(* Logix 5000 project; controller FV vendor 1 type 14 code 217 rev 31.11; software revision 31.00; part 26 of 63 *)
(* tags used below, declared in another part *)
   Alarm_Reset : BOOL;
   CheckTimeMask : INT;
   comms_to_mc_write_enabled : BOOL;
   comms_to_mv_route_write_enabled : BOOL;
   Default_Check_Time : DINT;
   Delphi_Does_Eng_Func : BOOL;
   FR_B3 : INT[255];   // BINARY
   fr_comms_from_mv_route : MESSAGE;
   fr_comms_from_mvfv_cip : MESSAGE;
   fr_comms_to_MC : MESSAGE;
   fr_comms_to_MC_timer : TIMER;
   fr_comms_to_mv_route : MESSAGE;
   fr_comms_to_mv_route_timer : TIMER;
   FR_FV27_AV08 : PlantItem;   // FV27_AV08
   FR_FV28_AV08 : PlantItem;   // FV28_AV08
   FR_FV29_AV08 : PlantItem;   // FV29_AV08
   FR_FV30_AV08 : PlantItem;   // FV30_AV08
   FR_FV31_AV08 : PlantItem;   // FV31_AV08
   FR_FVR1_P01 : PlantItem;   // FVR1_P01
   FR_FVR1_P01_ALARM : ALARM_DIGITAL;
   FR_FVR1_P01_D : ALIAS FOR RIO_Rack_2:5:O.Data.5;
   FR_FVR1_P01_R : ALIAS FOR RIO_Rack_2:4:I.Data.9;
   FR_FVS_P01 : PlantItem;   // FVS_P01
   FR_FVS_P01_ALARM : ALARM_DIGITAL;
   FR_FVS_P01_D : ALIAS FOR RIO_Rack_2:5:O.Data.0;
   FR_FVS_P01_R : ALIAS FOR RIO_Rack_2:4:I.Data.0;
   FR_GBM_P01 : PlantItem;   // GBM_P01
   FR_GBM_P01_ALARM : ALARM_DIGITAL;
   FR_GBM_P01_D : ALIAS FOR RIO_Rack_2:5:O.Data.2;
   FR_GBM_P01_R : ALIAS FOR RIO_Rack_2:4:I.Data.2;
   FR_N10 : INT[265];   // FV_AGING Comms to FV Aging PL C
   FR_N13 : INT[265];   // MV_ROUTE Comms to MV Routing PLC
   FR_N14 : INT[265];   // MVFV CIP Comms to MVFV CIP Un it PLC
   FR_N225 : INT[265];   // Original N File From SLC, No Description Available
   FR_N226 : INT[265];   // Original N File From SLC, No Description Available
   FR_N255 : INT[265];   // CHECKWORDS
   FR_N99 : INT[265];   // COMMENT Comment Lines
   FR_T19 : TIMER[255];   // HEARTBEAT Heartbeat Timers
   FR_T4 : TIMER[255];   // TIMER
   FR_YM_P01 : PlantItem;   // YM_P01
   FR_YM_P01_ALARM : ALARM_DIGITAL;
   FR_YM_P01_D : ALIAS FOR RIO_Rack_2:5:O.Data.1;
   FR_YM_P01_R : ALIAS FOR RIO_Rack_2:4:I.Data.1;
   FR_YM_P01_T : ALIAS FOR RIO_Rack_2:4:I.Data.5;
   FR_YM_P02 : PlantItem;   // YM_P02
   FR_YM_P02_ALARM : ALARM_DIGITAL;
   FR_YM_P02_D : ALIAS FOR RIO_Rack_2:5:O.Data.3;
   FR_YM_P02_R : ALIAS FOR RIO_Rack_2:4:I.Data.3;
   FR_YM_P02_T : ALIAS FOR RIO_Rack_2:4:I.Data.7;
   FR_YM_P03 : PlantItem;   // YM_P03
   FR_YM_P03_ALARM : ALARM_DIGITAL;
   FR_YM_P03_D : ALIAS FOR RIO_Rack_2:5:O.Data.4;
   FR_YM_P03_R : ALIAS FOR RIO_Rack_2:4:I.Data.8;
   FR_YM_P03_T : ALIAS FOR RIO_Rack_2:4:I.Data.12;
   FV_N191 : INT[255];   // FVR COMMS
   Item_Faults_Are_Latched : BOOL;
   Item_Simulation_Flag : BOOL;
   One_Second_One_Scan : ALIAS FOR One_Second_1_scan;
   reset_msg_interval : BOOL;
   Scada_Pump_Fault_No : DINT;
   Scada_Pump_H_Fault_No : DINT;
   Scada_Pump_T_Fault_No : DINT;
   TempChecktime : DINT;
   Unused_Healthy_Feedback : BOOL;
   Unused_NotTripped_Feedback : BOOL;
(* FR_Common, continued *)

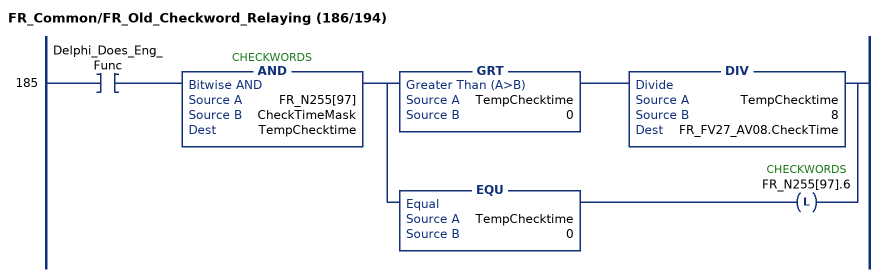
   [picture p490: FR_Common/FR_Old_Checkword_Relaying rungs 185-185]
   185: XIC(Delphi_Does_Eng_Func)AND(FR_N255[97],CheckTimeMask,TempChecktime)[GRT(TempChecktime,0) DIV(TempChecktime,8,FR_FV27_AV08.CheckTime) ,EQU(TempChecktime,0) OTL(FR_N255[97].6) ];
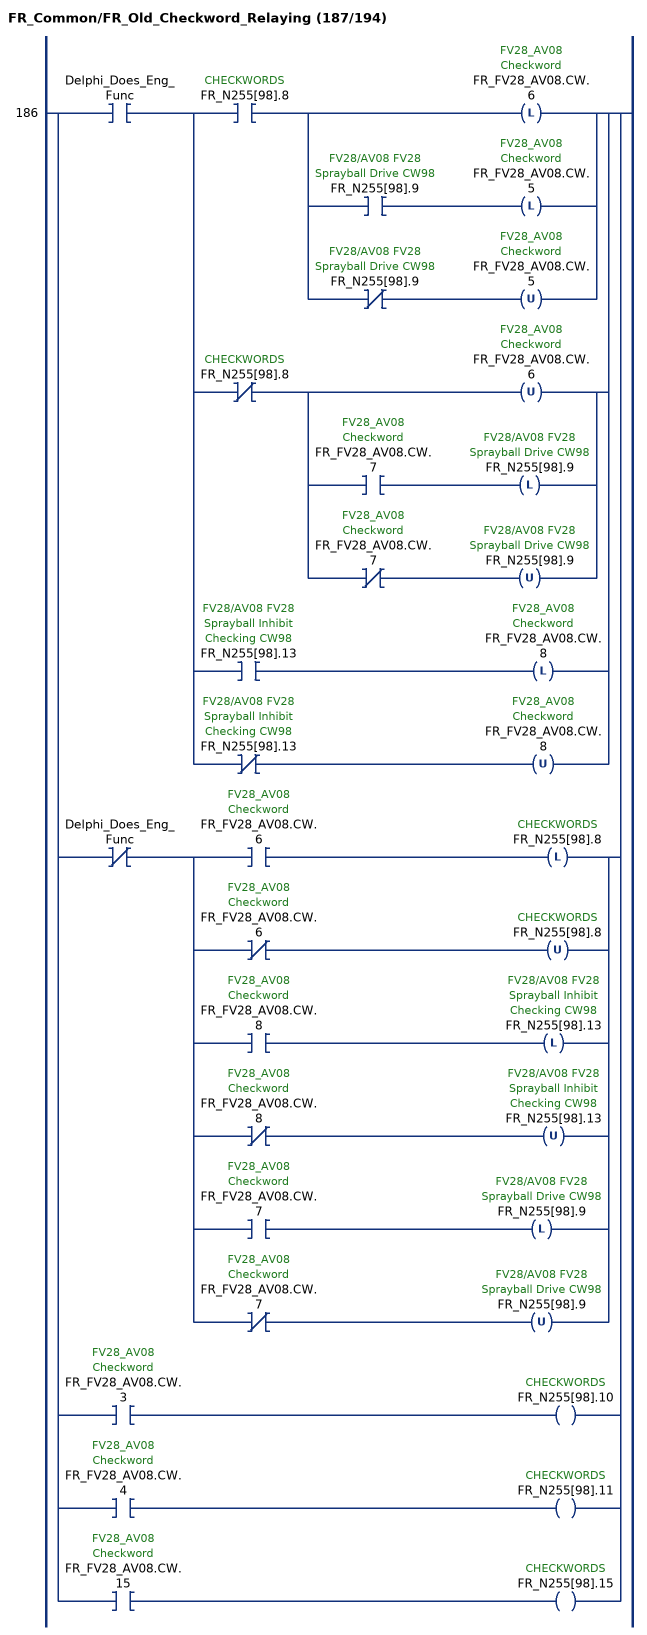
   186: [XIC(Delphi_Does_Eng_Func) [[XIC(FR_N255[98].8) [OTL(FR_FV28_AV08.CW.6) ,XIC(FR_N255[98].9) OTL(FR_FV28_AV08.CW.5) ,XIO(FR_N255[98].9) OTU(FR_FV28_AV08.CW.5) ] ,XIO(FR_N255[98].8) [OTU(FR_FV28_AV08.CW.6) ,[XIC(FR_FV28_AV08.CW.7) OTL(FR_N255[98].9) ,XIO(FR_FV28_AV08.CW.7) OTU(FR_N255[98].9) ] ] ] ,[XIC(FR_N255[98].13) OTL(FR_FV28_AV08.CW.8) ,XIO(FR_N255[98].13) OTU(FR_FV28_AV08.CW.8) ] ] ,XIO(Delphi_Does_Eng_Func) [[XIC(FR_FV28_AV08.CW.6) OTL(FR_N255[98].8) ,XIO(FR_FV28_AV08.CW.6) OTU(FR_N255[98].8) ] ,[XIC(FR_FV28_AV08.CW.8) OTL(FR_N255[98].13) ,XIO(FR_FV28_AV08.CW.8) OTU(FR_N255[98].13) ] ,[XIC(FR_FV28_AV08.CW.7) OTL(FR_N255[98].9) ,XIO(FR_FV28_AV08.CW.7) OTU(FR_N255[98].9) ] ] ,XIC(FR_FV28_AV08.CW.3) OTE(FR_N255[98].10) ,XIC(FR_FV28_AV08.CW.4) OTE(FR_N255[98].11) ,XIC(FR_FV28_AV08.CW.15) OTE(FR_N255[98].15) ];
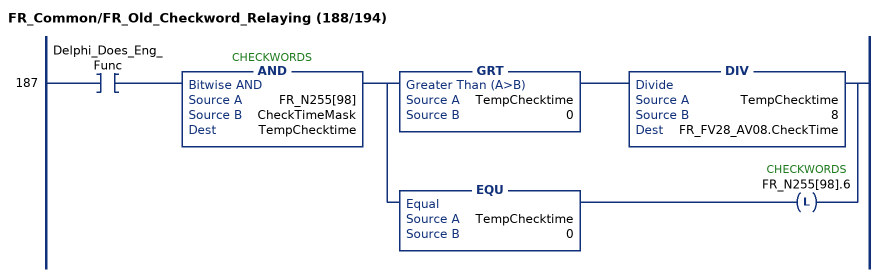
   187: XIC(Delphi_Does_Eng_Func)AND(FR_N255[98],CheckTimeMask,TempChecktime)[GRT(TempChecktime,0) DIV(TempChecktime,8,FR_FV28_AV08.CheckTime) ,EQU(TempChecktime,0) OTL(FR_N255[98].6) ];
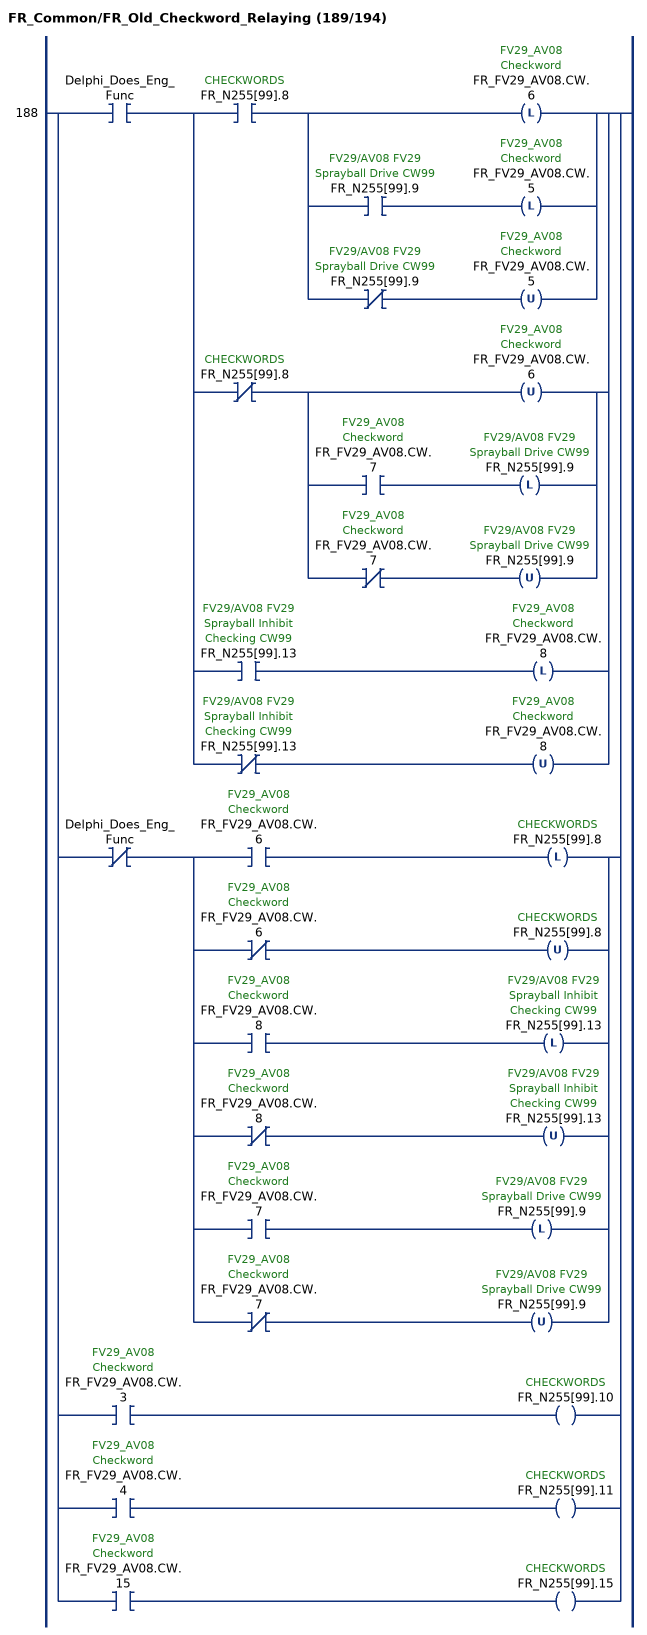
   188: [XIC(Delphi_Does_Eng_Func) [[XIC(FR_N255[99].8) [OTL(FR_FV29_AV08.CW.6) ,XIC(FR_N255[99].9) OTL(FR_FV29_AV08.CW.5) ,XIO(FR_N255[99].9) OTU(FR_FV29_AV08.CW.5) ] ,XIO(FR_N255[99].8) [OTU(FR_FV29_AV08.CW.6) ,[XIC(FR_FV29_AV08.CW.7) OTL(FR_N255[99].9) ,XIO(FR_FV29_AV08.CW.7) OTU(FR_N255[99].9) ] ] ] ,[XIC(FR_N255[99].13) OTL(FR_FV29_AV08.CW.8) ,XIO(FR_N255[99].13) OTU(FR_FV29_AV08.CW.8) ] ] ,XIO(Delphi_Does_Eng_Func) [[XIC(FR_FV29_AV08.CW.6) OTL(FR_N255[99].8) ,XIO(FR_FV29_AV08.CW.6) OTU(FR_N255[99].8) ] ,[XIC(FR_FV29_AV08.CW.8) OTL(FR_N255[99].13) ,XIO(FR_FV29_AV08.CW.8) OTU(FR_N255[99].13) ] ,[XIC(FR_FV29_AV08.CW.7) OTL(FR_N255[99].9) ,XIO(FR_FV29_AV08.CW.7) OTU(FR_N255[99].9) ] ] ,XIC(FR_FV29_AV08.CW.3) OTE(FR_N255[99].10) ,XIC(FR_FV29_AV08.CW.4) OTE(FR_N255[99].11) ,XIC(FR_FV29_AV08.CW.15) OTE(FR_N255[99].15) ];
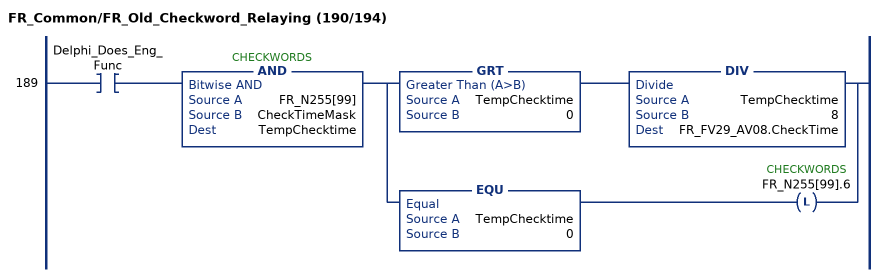
   189: XIC(Delphi_Does_Eng_Func)AND(FR_N255[99],CheckTimeMask,TempChecktime)[GRT(TempChecktime,0) DIV(TempChecktime,8,FR_FV29_AV08.CheckTime) ,EQU(TempChecktime,0) OTL(FR_N255[99].6) ];
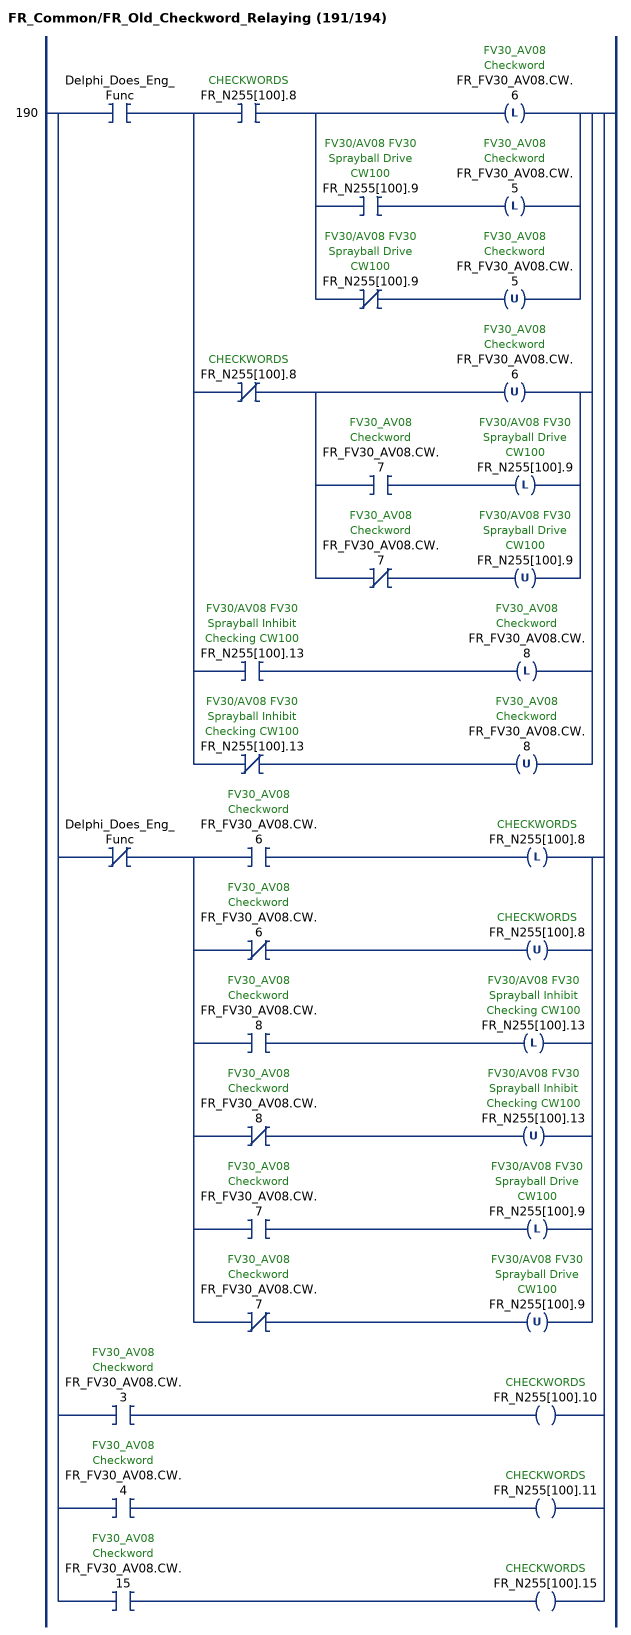
   190: [XIC(Delphi_Does_Eng_Func) [[XIC(FR_N255[100].8) [OTL(FR_FV30_AV08.CW.6) ,XIC(FR_N255[100].9) OTL(FR_FV30_AV08.CW.5) ,XIO(FR_N255[100].9) OTU(FR_FV30_AV08.CW.5) ] ,XIO(FR_N255[100].8) [OTU(FR_FV30_AV08.CW.6) ,[XIC(FR_FV30_AV08.CW.7) OTL(FR_N255[100].9) ,XIO(FR_FV30_AV08.CW.7) OTU(FR_N255[100].9) ] ] ] ,[XIC(FR_N255[100].13) OTL(FR_FV30_AV08.CW.8) ,XIO(FR_N255[100].13) OTU(FR_FV30_AV08.CW.8) ] ] ,XIO(Delphi_Does_Eng_Func) [[XIC(FR_FV30_AV08.CW.6) OTL(FR_N255[100].8) ,XIO(FR_FV30_AV08.CW.6) OTU(FR_N255[100].8) ] ,[XIC(FR_FV30_AV08.CW.8) OTL(FR_N255[100].13) ,XIO(FR_FV30_AV08.CW.8) OTU(FR_N255[100].13) ] ,[XIC(FR_FV30_AV08.CW.7) OTL(FR_N255[100].9) ,XIO(FR_FV30_AV08.CW.7) OTU(FR_N255[100].9) ] ] ,XIC(FR_FV30_AV08.CW.3) OTE(FR_N255[100].10) ,XIC(FR_FV30_AV08.CW.4) OTE(FR_N255[100].11) ,XIC(FR_FV30_AV08.CW.15) OTE(FR_N255[100].15) ];
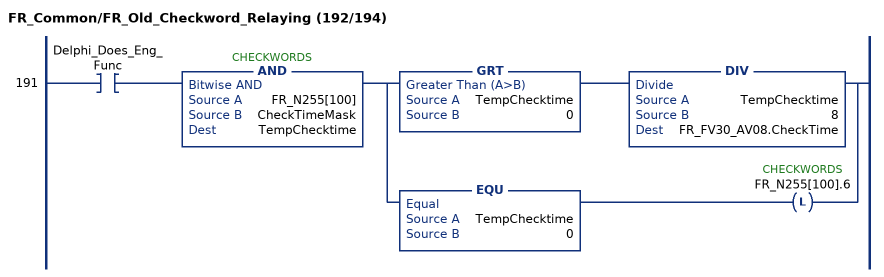
   191: XIC(Delphi_Does_Eng_Func)AND(FR_N255[100],CheckTimeMask,TempChecktime)[GRT(TempChecktime,0) DIV(TempChecktime,8,FR_FV30_AV08.CheckTime) ,EQU(TempChecktime,0) OTL(FR_N255[100].6) ];
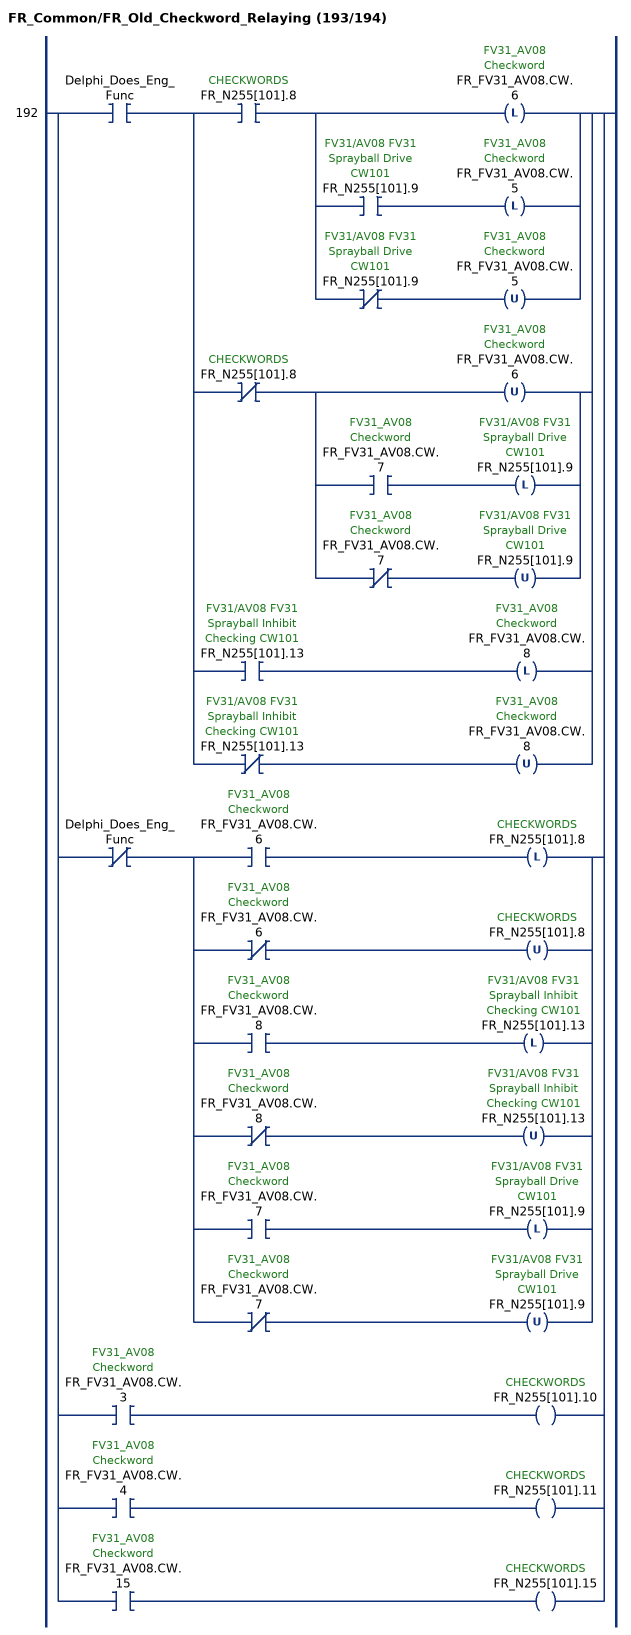
   192: [XIC(Delphi_Does_Eng_Func) [[XIC(FR_N255[101].8) [OTL(FR_FV31_AV08.CW.6) ,XIC(FR_N255[101].9) OTL(FR_FV31_AV08.CW.5) ,XIO(FR_N255[101].9) OTU(FR_FV31_AV08.CW.5) ] ,XIO(FR_N255[101].8) [OTU(FR_FV31_AV08.CW.6) ,[XIC(FR_FV31_AV08.CW.7) OTL(FR_N255[101].9) ,XIO(FR_FV31_AV08.CW.7) OTU(FR_N255[101].9) ] ] ] ,[XIC(FR_N255[101].13) OTL(FR_FV31_AV08.CW.8) ,XIO(FR_N255[101].13) OTU(FR_FV31_AV08.CW.8) ] ] ,XIO(Delphi_Does_Eng_Func) [[XIC(FR_FV31_AV08.CW.6) OTL(FR_N255[101].8) ,XIO(FR_FV31_AV08.CW.6) OTU(FR_N255[101].8) ] ,[XIC(FR_FV31_AV08.CW.8) OTL(FR_N255[101].13) ,XIO(FR_FV31_AV08.CW.8) OTU(FR_N255[101].13) ] ,[XIC(FR_FV31_AV08.CW.7) OTL(FR_N255[101].9) ,XIO(FR_FV31_AV08.CW.7) OTU(FR_N255[101].9) ] ] ,XIC(FR_FV31_AV08.CW.3) OTE(FR_N255[101].10) ,XIC(FR_FV31_AV08.CW.4) OTE(FR_N255[101].11) ,XIC(FR_FV31_AV08.CW.15) OTE(FR_N255[101].15) ];
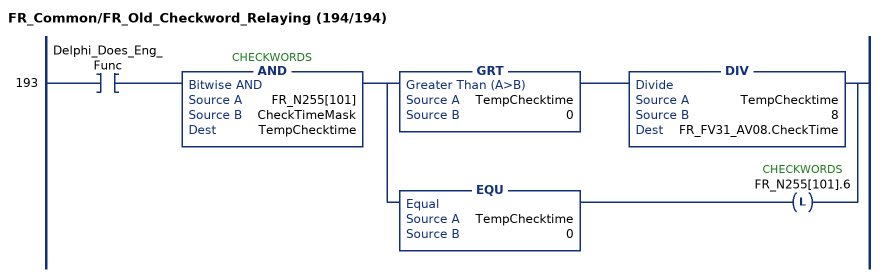
   193: XIC(Delphi_Does_Eng_Func)AND(FR_N255[101],CheckTimeMask,TempChecktime)[GRT(TempChecktime,0) DIV(TempChecktime,8,FR_FV31_AV08.CheckTime) ,EQU(TempChecktime,0) OTL(FR_N255[101].6) ];
END_ROUTINE

ROUTINE FR_PLC_COMMS_10   (* ladder *)
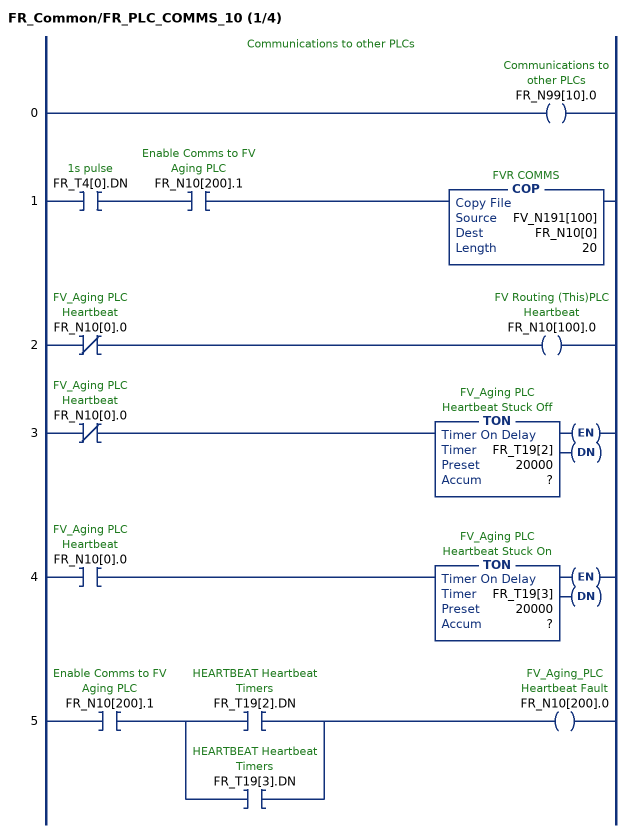
   // Communications to other PLCs
   0: OTE(FR_N99[10].0);
   1: XIC(FR_T4[0].DN)XIC(FR_N10[200].1)COP(FV_N191[100],FR_N10[0],20);
   2: XIO(FR_N10[0].0)OTE(FR_N10[100].0);
   3: XIO(FR_N10[0].0)TON(FR_T19[2],?,?);
   4: XIC(FR_N10[0].0)TON(FR_T19[3],?,?);
   5: XIC(FR_N10[200].1)[XIC(FR_T19[2].DN) ,XIC(FR_T19[3].DN) ]OTE(FR_N10[200].0);
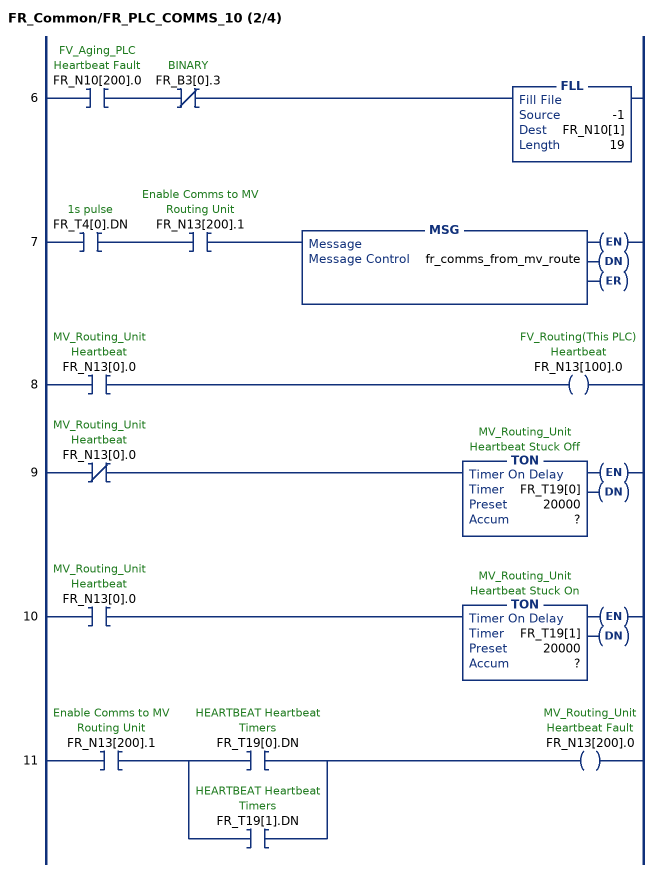
   6: XIC(FR_N10[200].0)XIO(FR_B3[0].3)FLL(-1,FR_N10[1],19);
   7: XIC(FR_T4[0].DN)XIC(FR_N13[200].1)MSG(fr_comms_from_mv_route);
   8: XIC(FR_N13[0].0)OTE(FR_N13[100].0);
   9: XIO(FR_N13[0].0)TON(FR_T19[0],?,?);
   10: XIC(FR_N13[0].0)TON(FR_T19[1],?,?);
   11: XIC(FR_N13[200].1)[XIC(FR_T19[0].DN) ,XIC(FR_T19[1].DN) ]OTE(FR_N13[200].0);
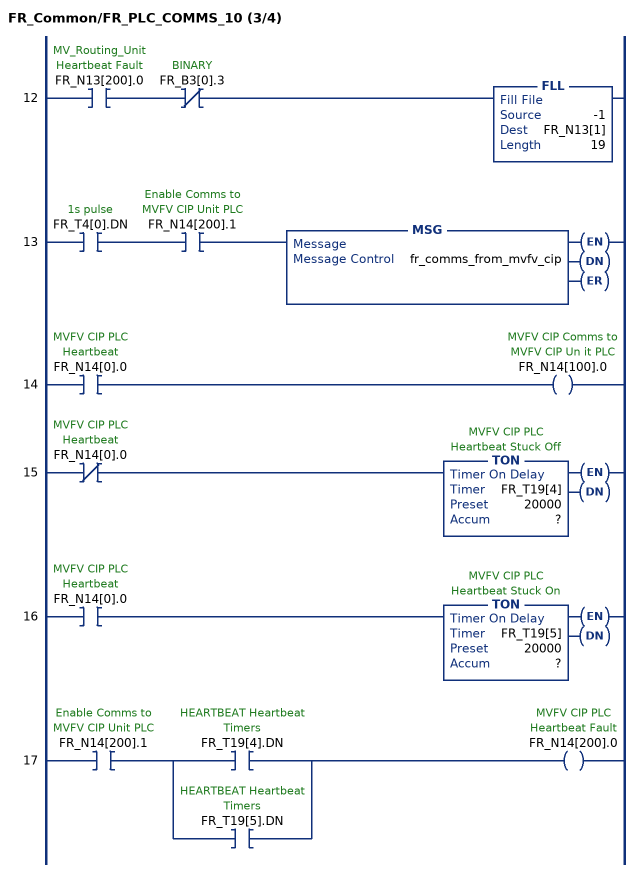
   12: XIC(FR_N13[200].0)XIO(FR_B3[0].3)FLL(-1,FR_N13[1],19);
   13: XIC(FR_T4[0].DN)XIC(FR_N14[200].1)MSG(fr_comms_from_mvfv_cip);
   14: XIC(FR_N14[0].0)OTE(FR_N14[100].0);
   15: XIO(FR_N14[0].0)TON(FR_T19[4],?,?);
   16: XIC(FR_N14[0].0)TON(FR_T19[5],?,?);
   17: XIC(FR_N14[200].1)[XIC(FR_T19[4].DN) ,XIC(FR_T19[5].DN) ]OTE(FR_N14[200].0);
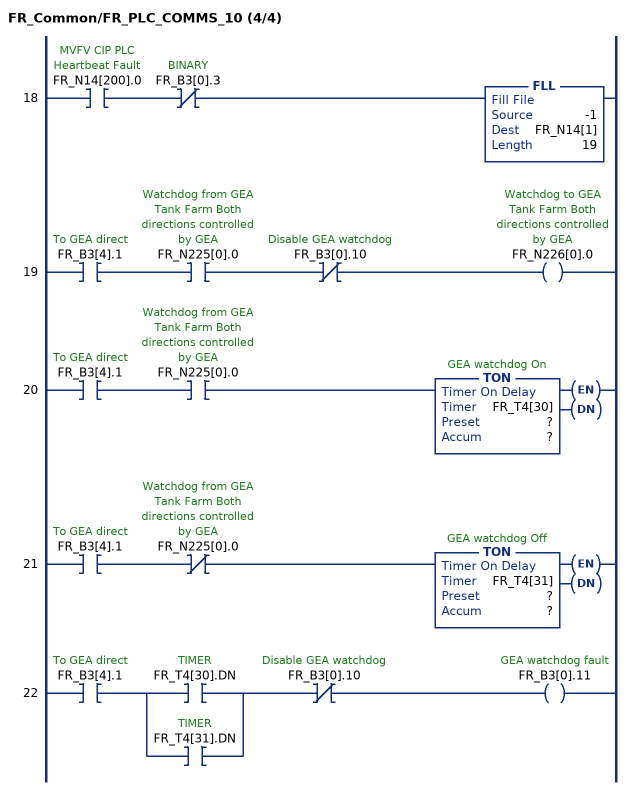
   18: XIC(FR_N14[200].0)XIO(FR_B3[0].3)FLL(-1,FR_N14[1],19);
   19: XIC(FR_B3[4].1)XIC(FR_N225[0].0)XIO(FR_B3[0].10)OTE(FR_N226[0].0);
   20: XIC(FR_B3[4].1)XIC(FR_N225[0].0)TON(FR_T4[30],?,?);
   21: XIC(FR_B3[4].1)XIO(FR_N225[0].0)TON(FR_T4[31],?,?);
   22: XIC(FR_B3[4].1)[XIC(FR_T4[30].DN) ,XIC(FR_T4[31].DN) ]XIO(FR_B3[0].10)OTE(FR_B3[0].11);
END_ROUTINE

ROUTINE FR_PLC_COMMS_Write_Replacements   (* ladder *)
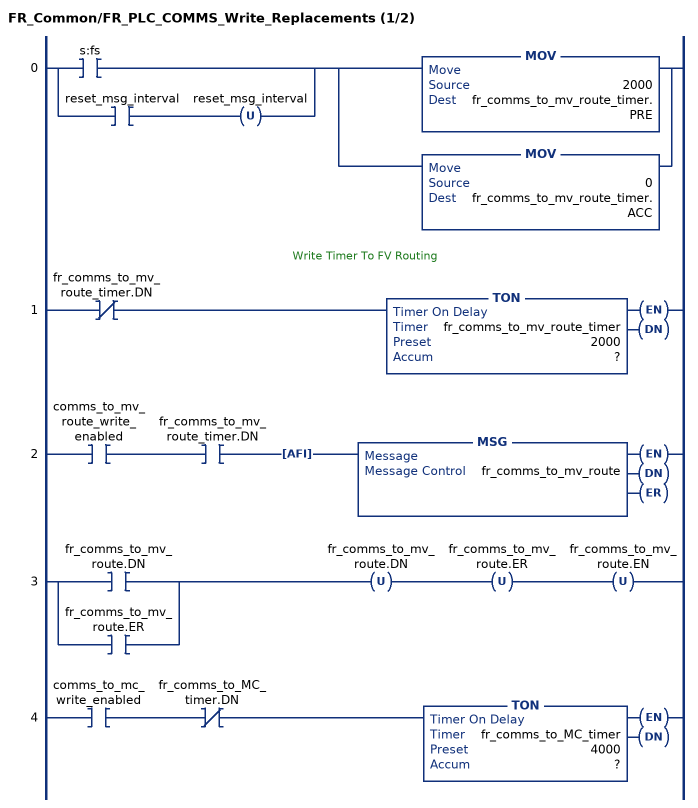
   0: [XIC(s:fs) ,XIC(reset_msg_interval) OTU(reset_msg_interval) ][MOV(2000,fr_comms_to_mv_route_timer.PRE) ,MOV(0,fr_comms_to_mv_route_timer.ACC) ];
   // Write Timer To FV Routing
   1: XIO(fr_comms_to_mv_route_timer.DN)TON(fr_comms_to_mv_route_timer,?,?);
   2: XIC(comms_to_mv_route_write_enabled)XIC(fr_comms_to_mv_route_timer.DN)AFI()MSG(fr_comms_to_mv_route);
   3: [XIC(fr_comms_to_mv_route.DN) ,XIC(fr_comms_to_mv_route.ER) ]OTU(fr_comms_to_mv_route.DN)OTU(fr_comms_to_mv_route.ER)OTU(fr_comms_to_mv_route.EN);
   4: XIC(comms_to_mc_write_enabled)XIO(fr_comms_to_MC_timer.DN)TON(fr_comms_to_MC_timer,?,?);
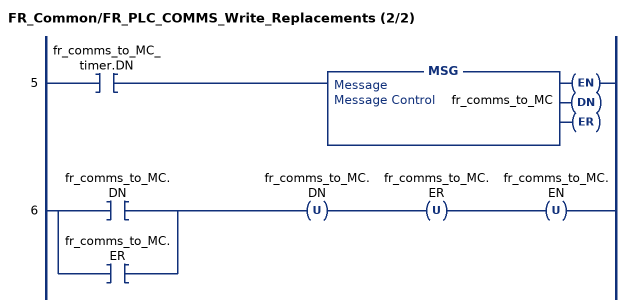
   5: XIC(fr_comms_to_MC_timer.DN)MSG(fr_comms_to_MC);
   6: [XIC(fr_comms_to_MC.DN) ,XIC(fr_comms_to_MC.ER) ]OTU(fr_comms_to_MC.DN)OTU(fr_comms_to_MC.ER)OTU(fr_comms_to_MC.EN);
END_ROUTINE

ROUTINE FR_Pumps   (* ladder *)
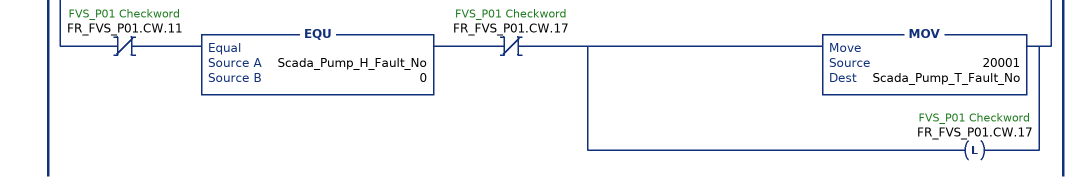
   0: [NEQ(FR_FVS_P01.DriveBits,0) OTE(FR_FVS_P01.CW.0) ,[XIC(FR_FVS_P01.CW.0) XIO(FR_FVS_P01.CW.6) ,XIC(FR_FVS_P01.CW.5) XIC(FR_FVS_P01.CW.6) ] OTE(FR_FVS_P01.CW.7) ,XIC(FR_FVS_P01.CW.7) OTE(FR_FVS_P01_D) ,XIC(S:FS) [OTU(FR_FVS_P01.CW.6) ,LEQ(FR_FVS_P01.CheckTime,0) MOV(Default_Check_Time,FR_FVS_P01.CheckTime) ] ,[[XIC(FR_FVS_P01_R) XIO(Item_Simulation_Flag) ,XIC(Item_Simulation_Flag) [XIC(FR_FVS_P01.CW.7) XIO(FR_FVS_P01.CW.2) ,XIO(FR_FVS_P01.CW.7) XIC(FR_FVS_P01.CW.2) ] ] OTE(FR_FVS_P01.CW.3) ,[XIC(Item_Simulation_Flag) ,XIC(FR_FVS_P01.CW.8) ,XIC(Unused_Healthy_Feedback) ] OTE(FR_FVS_P01.CW.10) ,[XIC(Item_Simulation_Flag) ,XIC(FR_FVS_P01.CW.8) ,XIC(Unused_NotTripped_Feedback) ] OTE(FR_FVS_P01.CW.11) ] ,[XIC(FR_FVS_P01.CW.7) XIO(FR_FVS_P01.CW.1) ,XIO(FR_FVS_P01.CW.7) XIC(FR_FVS_P01.CW.1) ] CLR(FR_FVS_P01.CheckTimer) ,XIC(One_Second_One_Scan) LES(FR_FVS_P01.CheckTimer,FR_FVS_P01.CheckTime) ADD(FR_FVS_P01.CheckTimer,1,FR_FVS_P01.CheckTimer) ,XIO(FR_FVS_P01.CW.15) OTU(FR_FVS_P01.CW.14) ,[GEQ(FR_FVS_P01.CheckTimer,FR_FVS_P01.CheckTime) [XIC(FR_FVS_P01.CW.7) XIO(FR_FVS_P01.CW.3) ,XIO(FR_FVS_P01.CW.7) XIC(FR_FVS_P01.CW.3) ] ,XIO(FR_FVS_P01.CW.10) ,XIO(FR_FVS_P01.CW.11) ,XIC(FR_FVS_P01.CW.15) XIC(Item_Faults_Are_Latched) ,XIC(FR_FVS_P01.CW.9) ] XIO(FR_FVS_P01.CW.8) XIO(Alarm_Reset) [OTE(FR_FVS_P01.CW.15) ,ALMD(FR_FVS_P01_ALARM,0,0,0,0) ] ,XIC(FR_FVS_P01.CW.7) OTE(FR_FVS_P01.CW.1) ,XIC(FR_FVS_P01.CW.15) EQU(Scada_Pump_Fault_No,0) XIO(FR_FVS_P01.CW.14) [MOV(20001,Scada_Pump_Fault_No) ,OTL(FR_FVS_P01.CW.14) ] ,XIO(FR_FVS_P01.CW.10) EQU(Scada_Pump_H_Fault_No,0) XIO(FR_FVS_P01.CW.16) [MOV(20001,Scada_Pump_H_Fault_No) ,OTL(FR_FVS_P01.CW.16) ] ,XIO(FR_FVS_P01.CW.11) EQU(Scada_Pump_H_Fault_No,0) XIO(FR_FVS_P01.CW.17) [MOV(20001,Scada_Pump_T_Fault_No) ,OTL(FR_FVS_P01.CW.17) ] ];
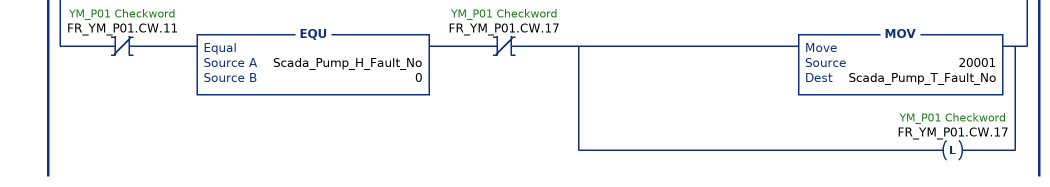
   1: [NEQ(FR_YM_P01.DriveBits,0) OTE(FR_YM_P01.CW.0) ,[XIC(FR_YM_P01.CW.0) XIO(FR_YM_P01.CW.6) ,XIC(FR_YM_P01.CW.5) XIC(FR_YM_P01.CW.6) ] OTE(FR_YM_P01.CW.7) ,XIC(FR_YM_P01.CW.7) OTE(FR_YM_P01_D) ,XIC(S:FS) [OTU(FR_YM_P01.CW.6) ,LEQ(FR_YM_P01.CheckTime,0) MOV(Default_Check_Time,FR_YM_P01.CheckTime) ] ,[[XIC(FR_YM_P01_R) XIO(Item_Simulation_Flag) ,XIC(Item_Simulation_Flag) [XIC(FR_YM_P01.CW.7) XIO(FR_YM_P01.CW.2) ,XIO(FR_YM_P01.CW.7) XIC(FR_YM_P01.CW.2) ] ] OTE(FR_YM_P01.CW.3) ,[XIC(Item_Simulation_Flag) ,XIC(FR_YM_P01.CW.8) ,XIC(Unused_Healthy_Feedback) ] OTE(FR_YM_P01.CW.10) ,[XIC(Item_Simulation_Flag) ,XIC(FR_YM_P01.CW.8) ,XIO(FR_YM_P01_T) ] OTE(FR_YM_P01.CW.11) ] ,[XIC(FR_YM_P01.CW.7) XIO(FR_YM_P01.CW.1) ,XIO(FR_YM_P01.CW.7) XIC(FR_YM_P01.CW.1) ] CLR(FR_YM_P01.CheckTimer) ,XIC(One_Second_One_Scan) LES(FR_YM_P01.CheckTimer,FR_YM_P01.CheckTime) ADD(FR_YM_P01.CheckTimer,1,FR_YM_P01.CheckTimer) ,XIO(FR_YM_P01.CW.15) OTU(FR_YM_P01.CW.14) ,[GEQ(FR_YM_P01.CheckTimer,FR_YM_P01.CheckTime) [XIC(FR_YM_P01.CW.7) XIO(FR_YM_P01.CW.3) ,XIO(FR_YM_P01.CW.7) XIC(FR_YM_P01.CW.3) ] ,XIO(FR_YM_P01.CW.10) ,XIO(FR_YM_P01.CW.11) ,XIC(FR_YM_P01.CW.15) XIC(Item_Faults_Are_Latched) ,XIC(FR_YM_P01.CW.9) ] XIO(FR_YM_P01.CW.8) XIO(Alarm_Reset) [OTE(FR_YM_P01.CW.15) ,ALMD(FR_YM_P01_ALARM,0,0,0,0) ] ,XIC(FR_YM_P01.CW.7) OTE(FR_YM_P01.CW.1) ,XIC(FR_YM_P01.CW.15) EQU(Scada_Pump_Fault_No,0) XIO(FR_YM_P01.CW.14) [MOV(20001,Scada_Pump_Fault_No) ,OTL(FR_YM_P01.CW.14) ] ,XIO(FR_YM_P01.CW.10) EQU(Scada_Pump_H_Fault_No,0) XIO(FR_YM_P01.CW.16) [MOV(20001,Scada_Pump_H_Fault_No) ,OTL(FR_YM_P01.CW.16) ] ,XIO(FR_YM_P01.CW.11) EQU(Scada_Pump_H_Fault_No,0) XIO(FR_YM_P01.CW.17) [MOV(20001,Scada_Pump_T_Fault_No) ,OTL(FR_YM_P01.CW.17) ] ];
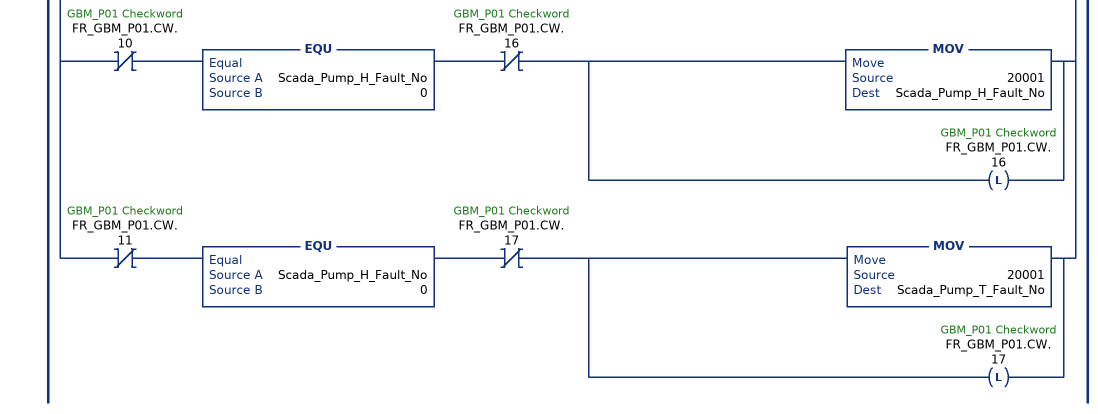
   2: [NEQ(FR_GBM_P01.DriveBits,0) OTE(FR_GBM_P01.CW.0) ,[XIC(FR_GBM_P01.CW.0) XIO(FR_GBM_P01.CW.6) ,XIC(FR_GBM_P01.CW.5) XIC(FR_GBM_P01.CW.6) ] OTE(FR_GBM_P01.CW.7) ,XIC(FR_GBM_P01.CW.7) OTE(FR_GBM_P01_D) ,XIC(S:FS) [OTU(FR_GBM_P01.CW.6) ,LEQ(FR_GBM_P01.CheckTime,0) MOV(Default_Check_Time,FR_GBM_P01.CheckTime) ] ,[[XIC(FR_GBM_P01_R) XIO(Item_Simulation_Flag) ,XIC(Item_Simulation_Flag) [XIC(FR_GBM_P01.CW.7) XIO(FR_GBM_P01.CW.2) ,XIO(FR_GBM_P01.CW.7) XIC(FR_GBM_P01.CW.2) ] ] OTE(FR_GBM_P01.CW.3) ,[XIC(Item_Simulation_Flag) ,XIC(FR_GBM_P01.CW.8) ,XIC(Unused_Healthy_Feedback) ] OTE(FR_GBM_P01.CW.10) ,[XIC(Item_Simulation_Flag) ,XIC(FR_GBM_P01.CW.8) ,XIC(Unused_NotTripped_Feedback) ] OTE(FR_GBM_P01.CW.11) ] ,[XIC(FR_GBM_P01.CW.7) XIO(FR_GBM_P01.CW.1) ,XIO(FR_GBM_P01.CW.7) XIC(FR_GBM_P01.CW.1) ] CLR(FR_GBM_P01.CheckTimer) ,XIC(One_Second_One_Scan) LES(FR_GBM_P01.CheckTimer,FR_GBM_P01.CheckTime) ADD(FR_GBM_P01.CheckTimer,1,FR_GBM_P01.CheckTimer) ,XIO(FR_GBM_P01.CW.15) OTU(FR_GBM_P01.CW.14) ,[GEQ(FR_GBM_P01.CheckTimer,FR_GBM_P01.CheckTime) [XIC(FR_GBM_P01.CW.7) XIO(FR_GBM_P01.CW.3) ,XIO(FR_GBM_P01.CW.7) XIC(FR_GBM_P01.CW.3) ] ,XIO(FR_GBM_P01.CW.10) ,XIO(FR_GBM_P01.CW.11) ,XIC(FR_GBM_P01.CW.15) XIC(Item_Faults_Are_Latched) ,XIC(FR_GBM_P01.CW.9) ] XIO(FR_GBM_P01.CW.8) XIO(Alarm_Reset) [OTE(FR_GBM_P01.CW.15) ,ALMD(FR_GBM_P01_ALARM,0,0,0,0) ] ,XIC(FR_GBM_P01.CW.7) OTE(FR_GBM_P01.CW.1) ,XIC(FR_GBM_P01.CW.15) EQU(Scada_Pump_Fault_No,0) XIO(FR_GBM_P01.CW.14) [MOV(20001,Scada_Pump_Fault_No) ,OTL(FR_GBM_P01.CW.14) ] ,XIO(FR_GBM_P01.CW.10) EQU(Scada_Pump_H_Fault_No,0) XIO(FR_GBM_P01.CW.16) [MOV(20001,Scada_Pump_H_Fault_No) ,OTL(FR_GBM_P01.CW.16) ] ,XIO(FR_GBM_P01.CW.11) EQU(Scada_Pump_H_Fault_No,0) XIO(FR_GBM_P01.CW.17) [MOV(20001,Scada_Pump_T_Fault_No) ,OTL(FR_GBM_P01.CW.17) ] ];
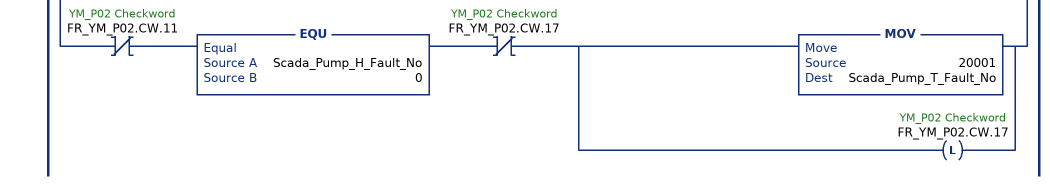
   3: [NEQ(FR_YM_P02.DriveBits,0) OTE(FR_YM_P02.CW.0) ,[XIC(FR_YM_P02.CW.0) XIO(FR_YM_P02.CW.6) ,XIC(FR_YM_P02.CW.5) XIC(FR_YM_P02.CW.6) ] OTE(FR_YM_P02.CW.7) ,XIC(FR_YM_P02.CW.7) OTE(FR_YM_P02_D) ,XIC(S:FS) [OTU(FR_YM_P02.CW.6) ,LEQ(FR_YM_P02.CheckTime,0) MOV(Default_Check_Time,FR_YM_P02.CheckTime) ] ,[[XIC(FR_YM_P02_R) XIO(Item_Simulation_Flag) ,XIC(Item_Simulation_Flag) [XIC(FR_YM_P02.CW.7) XIO(FR_YM_P02.CW.2) ,XIO(FR_YM_P02.CW.7) XIC(FR_YM_P02.CW.2) ] ] OTE(FR_YM_P02.CW.3) ,[XIC(Item_Simulation_Flag) ,XIC(FR_YM_P02.CW.8) ,XIC(Unused_Healthy_Feedback) ] OTE(FR_YM_P02.CW.10) ,[XIC(Item_Simulation_Flag) ,XIC(FR_YM_P02.CW.8) ,XIO(FR_YM_P02_T) ] OTE(FR_YM_P02.CW.11) ] ,[XIC(FR_YM_P02.CW.7) XIO(FR_YM_P02.CW.1) ,XIO(FR_YM_P02.CW.7) XIC(FR_YM_P02.CW.1) ] CLR(FR_YM_P02.CheckTimer) ,XIC(One_Second_One_Scan) LES(FR_YM_P02.CheckTimer,FR_YM_P02.CheckTime) ADD(FR_YM_P02.CheckTimer,1,FR_YM_P02.CheckTimer) ,XIO(FR_YM_P02.CW.15) OTU(FR_YM_P02.CW.14) ,[GEQ(FR_YM_P02.CheckTimer,FR_YM_P02.CheckTime) [XIC(FR_YM_P02.CW.7) XIO(FR_YM_P02.CW.3) ,XIO(FR_YM_P02.CW.7) XIC(FR_YM_P02.CW.3) ] ,XIO(FR_YM_P02.CW.10) ,XIO(FR_YM_P02.CW.11) ,XIC(FR_YM_P02.CW.15) XIC(Item_Faults_Are_Latched) ,XIC(FR_YM_P02.CW.9) ] XIO(FR_YM_P02.CW.8) XIO(Alarm_Reset) [OTE(FR_YM_P02.CW.15) ,ALMD(FR_YM_P02_ALARM,0,0,0,0) ] ,XIC(FR_YM_P02.CW.7) OTE(FR_YM_P02.CW.1) ,XIC(FR_YM_P02.CW.15) EQU(Scada_Pump_Fault_No,0) XIO(FR_YM_P02.CW.14) [MOV(20001,Scada_Pump_Fault_No) ,OTL(FR_YM_P02.CW.14) ] ,XIO(FR_YM_P02.CW.10) EQU(Scada_Pump_H_Fault_No,0) XIO(FR_YM_P02.CW.16) [MOV(20001,Scada_Pump_H_Fault_No) ,OTL(FR_YM_P02.CW.16) ] ,XIO(FR_YM_P02.CW.11) EQU(Scada_Pump_H_Fault_No,0) XIO(FR_YM_P02.CW.17) [MOV(20001,Scada_Pump_T_Fault_No) ,OTL(FR_YM_P02.CW.17) ] ];
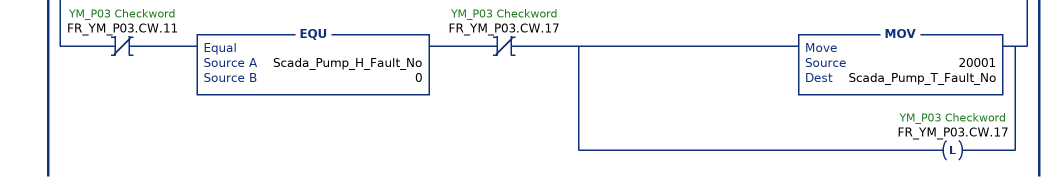
   4: [NEQ(FR_YM_P03.DriveBits,0) OTE(FR_YM_P03.CW.0) ,[XIC(FR_YM_P03.CW.0) XIO(FR_YM_P03.CW.6) ,XIC(FR_YM_P03.CW.5) XIC(FR_YM_P03.CW.6) ] OTE(FR_YM_P03.CW.7) ,XIC(FR_YM_P03.CW.7) OTE(FR_YM_P03_D) ,XIC(S:FS) [OTU(FR_YM_P03.CW.6) ,LEQ(FR_YM_P03.CheckTime,0) MOV(Default_Check_Time,FR_YM_P03.CheckTime) ] ,[[XIC(FR_YM_P03_R) XIO(Item_Simulation_Flag) ,XIC(Item_Simulation_Flag) [XIC(FR_YM_P03.CW.7) XIO(FR_YM_P03.CW.2) ,XIO(FR_YM_P03.CW.7) XIC(FR_YM_P03.CW.2) ] ] OTE(FR_YM_P03.CW.3) ,[XIC(Item_Simulation_Flag) ,XIC(FR_YM_P03.CW.8) ,XIC(Unused_Healthy_Feedback) ] OTE(FR_YM_P03.CW.10) ,[XIC(Item_Simulation_Flag) ,XIC(FR_YM_P03.CW.8) ,XIO(FR_YM_P03_T) ] OTE(FR_YM_P03.CW.11) ] ,[XIC(FR_YM_P03.CW.7) XIO(FR_YM_P03.CW.1) ,XIO(FR_YM_P03.CW.7) XIC(FR_YM_P03.CW.1) ] CLR(FR_YM_P03.CheckTimer) ,XIC(One_Second_One_Scan) LES(FR_YM_P03.CheckTimer,FR_YM_P03.CheckTime) ADD(FR_YM_P03.CheckTimer,1,FR_YM_P03.CheckTimer) ,XIO(FR_YM_P03.CW.15) OTU(FR_YM_P03.CW.14) ,[GEQ(FR_YM_P03.CheckTimer,FR_YM_P03.CheckTime) [XIC(FR_YM_P03.CW.7) XIO(FR_YM_P03.CW.3) ,XIO(FR_YM_P03.CW.7) XIC(FR_YM_P03.CW.3) ] ,XIO(FR_YM_P03.CW.10) ,XIO(FR_YM_P03.CW.11) ,XIC(FR_YM_P03.CW.15) XIC(Item_Faults_Are_Latched) ,XIC(FR_YM_P03.CW.9) ] XIO(FR_YM_P03.CW.8) XIO(Alarm_Reset) [OTE(FR_YM_P03.CW.15) ,ALMD(FR_YM_P03_ALARM,0,0,0,0) ] ,XIC(FR_YM_P03.CW.7) OTE(FR_YM_P03.CW.1) ,XIC(FR_YM_P03.CW.15) EQU(Scada_Pump_Fault_No,0) XIO(FR_YM_P03.CW.14) [MOV(20001,Scada_Pump_Fault_No) ,OTL(FR_YM_P03.CW.14) ] ,XIO(FR_YM_P03.CW.10) EQU(Scada_Pump_H_Fault_No,0) XIO(FR_YM_P03.CW.16) [MOV(20001,Scada_Pump_H_Fault_No) ,OTL(FR_YM_P03.CW.16) ] ,XIO(FR_YM_P03.CW.11) EQU(Scada_Pump_H_Fault_No,0) XIO(FR_YM_P03.CW.17) [MOV(20001,Scada_Pump_T_Fault_No) ,OTL(FR_YM_P03.CW.17) ] ];
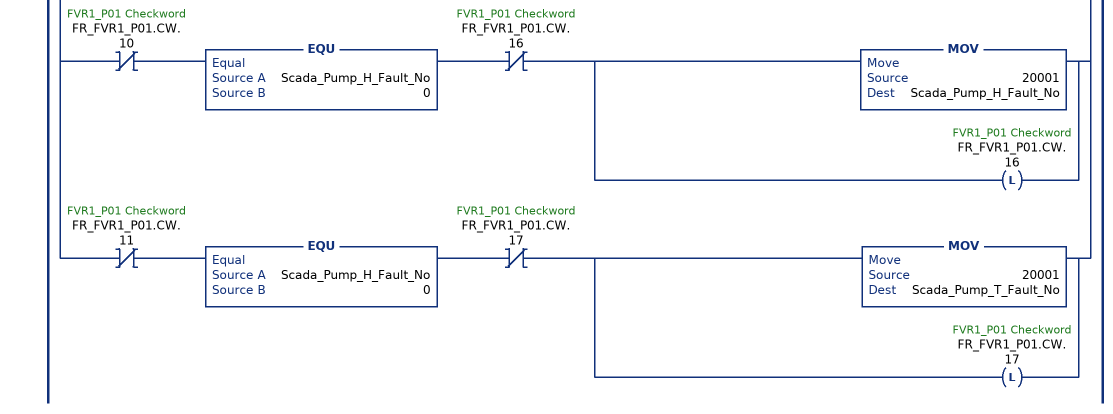
   5: [NEQ(FR_FVR1_P01.DriveBits,0) OTE(FR_FVR1_P01.CW.0) ,[XIC(FR_FVR1_P01.CW.0) XIO(FR_FVR1_P01.CW.6) ,XIC(FR_FVR1_P01.CW.5) XIC(FR_FVR1_P01.CW.6) ] OTE(FR_FVR1_P01.CW.7) ,XIC(FR_FVR1_P01.CW.7) OTE(FR_FVR1_P01_D) ,XIC(S:FS) [OTU(FR_FVR1_P01.CW.6) ,LEQ(FR_FVR1_P01.CheckTime,0) MOV(Default_Check_Time,FR_FVR1_P01.CheckTime) ] ,[[XIC(FR_FVR1_P01_R) XIO(Item_Simulation_Flag) ,XIC(Item_Simulation_Flag) [XIC(FR_FVR1_P01.CW.7) XIO(FR_FVR1_P01.CW.2) ,XIO(FR_FVR1_P01.CW.7) XIC(FR_FVR1_P01.CW.2) ] ] OTE(FR_FVR1_P01.CW.3) ,[XIC(Item_Simulation_Flag) ,XIC(FR_FVR1_P01.CW.8) ,XIC(Unused_Healthy_Feedback) ] OTE(FR_FVR1_P01.CW.10) ,[XIC(Item_Simulation_Flag) ,XIC(FR_FVR1_P01.CW.8) ,XIC(Unused_NotTripped_Feedback) ] OTE(FR_FVR1_P01.CW.11) ] ,[XIC(FR_FVR1_P01.CW.7) XIO(FR_FVR1_P01.CW.1) ,XIO(FR_FVR1_P01.CW.7) XIC(FR_FVR1_P01.CW.1) ] CLR(FR_FVR1_P01.CheckTimer) ,XIC(One_Second_One_Scan) LES(FR_FVR1_P01.CheckTimer,FR_FVR1_P01.CheckTime) ADD(FR_FVR1_P01.CheckTimer,1,FR_FVR1_P01.CheckTimer) ,XIO(FR_FVR1_P01.CW.15) OTU(FR_FVR1_P01.CW.14) ,[GEQ(FR_FVR1_P01.CheckTimer,FR_FVR1_P01.CheckTime) [XIC(FR_FVR1_P01.CW.7) XIO(FR_FVR1_P01.CW.3) ,XIO(FR_FVR1_P01.CW.7) XIC(FR_FVR1_P01.CW.3) ] ,XIO(FR_FVR1_P01.CW.10) ,XIO(FR_FVR1_P01.CW.11) ,XIC(FR_FVR1_P01.CW.15) XIC(Item_Faults_Are_Latched) ,XIC(FR_FVR1_P01.CW.9) ] XIO(FR_FVR1_P01.CW.8) XIO(Alarm_Reset) [OTE(FR_FVR1_P01.CW.15) ,ALMD(FR_FVR1_P01_ALARM,0,0,0,0) ] ,XIC(FR_FVR1_P01.CW.7) OTE(FR_FVR1_P01.CW.1) ,XIC(FR_FVR1_P01.CW.15) EQU(Scada_Pump_Fault_No,0) XIO(FR_FVR1_P01.CW.14) [MOV(20001,Scada_Pump_Fault_No) ,OTL(FR_FVR1_P01.CW.14) ] ,XIO(FR_FVR1_P01.CW.10) EQU(Scada_Pump_H_Fault_No,0) XIO(FR_FVR1_P01.CW.16) [MOV(20001,Scada_Pump_H_Fault_No) ,OTL(FR_FVR1_P01.CW.16) ] ,XIO(FR_FVR1_P01.CW.11) EQU(Scada_Pump_H_Fault_No,0) XIO(FR_FVR1_P01.CW.17) [MOV(20001,Scada_Pump_T_Fault_No) ,OTL(FR_FVR1_P01.CW.17) ] ];
END_ROUTINE
